HMI tags "BWTS_BTCS"
   "80_From_HMI_RUN_BTCS" : Bool = PLC "80_From_HMI".RUN_BTCS, 1 s
   "80_From_HMI_RUN_BWTS" : Bool = PLC "80_From_HMI".RUN_BWTS, 1 s
   "2110_BTCS_CNTRL_DB_PRE_DWELL_HRS" : Int = PLC "2110_BTCS_CNTRL_DB".PRE_DWELL_HRS, 1 s
   "2110_BTCS_CNTRL_DB_DE_OX_HRS" : Int = PLC "80_From_HMI".MAN_AQ_INC_96, 1 s
   "2110_BTCS_CNTRL_DB_DE_OX_SP_HRS" : Int = PLC "2110_BTCS_CNTRL_DB".DE_OX_SP_HRS, 1 s
   "2110_BTCS_CNTRL_DB_DWELL_HRS" : Int = PLC "2110_BTCS_CNTRL_DB".DWELL_HRS, 1 s
   "2110_BTCS_CNTRL_DB_RE_OX_HRS" : Int = PLC "2110_BTCS_CNTRL_DB".RE_OX_HRS, 1 s
   "2110_BTCS_CNTRL_DB_RE_OX_SP_HRS" : Int = PLC "2110_BTCS_CNTRL_DB".RE_OX_SP_HRS, 1 s
   "2110_BTCS_CNTRL_DB_POST_DWELL_HRS" : Int = PLC "2110_BTCS_CNTRL_DB".POST_DWELL_HRS, 1 s
   "2110_BTCS_CNTRL_DB_PRE_DWELL_MINS" : Int = PLC "2110_BTCS_CNTRL_DB".PRE_DWELL_MINS, 1 s
   "2110_BTCS_CNTRL_DB_DE_OX_MINS" : Int = PLC "2110_BTCS_CNTRL_DB".DE_OX_MINS, 1 s
   "2110_BTCS_CNTRL_DB_DE_OX_SP_MINS" : Int = PLC "2110_BTCS_CNTRL_DB".DE_OX_SP_MINS, 1 s
   "2110_BTCS_CNTRL_DB_DWELL_MINS" : Int = PLC "2110_BTCS_CNTRL_DB".DWELL_MINS, 1 s
   "2110_BTCS_CNTRL_DB_RE_OX_MINS" : Int = PLC "2110_BTCS_CNTRL_DB".RE_OX_MINS, 1 s
   "2110_BTCS_CNTRL_DB_RE_OX_SP_MINS" : Int = PLC "2110_BTCS_CNTRL_DB".RE_OX_SP_MINS, 1 s
   "2110_BTCS_CNTRL_DB_POST_DWELL_MINS" : Int = PLC "2110_BTCS_CNTRL_DB".POST_DWELL_MINS, 1 s
   "2110_BTCS_CNTRL_DB_TOT_SEQ_HRS" : Int = PLC "2110_BTCS_CNTRL_DB".TOT_SEQ_HRS, 1 s
   "2110_BTCS_CNTRL_DB_TOT_SEQ_MINS" : Int = PLC "2110_BTCS_CNTRL_DB".TOT_SEQ_MINS, 1 s
   "2110_BTCS_CNTRL_DB_RMNG_SEQ_HRS" : Int = PLC "84_Setpoints".PIT358_InitialFill_Low, 1 s
   "2110_BTCS_CNTRL_DB_RMNG_SEQ_MINS" : Int = PLC "2110_BTCS_CNTRL_DB".RMNG_SEQ_MINS, 1 s
   "2110_BTCS_CNTRL_DB_BTCS_STATE" : Int = PLC "2110_BTCS_CNTRL_DB".BTCS_STATE, 1 s
   "2110_BTCS_CNTRL_DB_BTCS_STEP" : Int = PLC "2110_BTCS_CNTRL_DB".BTCS_STEP, 1 s
   "2110_BTCS_CNTRL_DB_START_SEQ" : Bool = PLC "2110_BTCS_CNTRL_DB".START_SEQ, 1 s
   "2110_BTCS_CNTRL_DB_STOP_SEQ" : Bool = PLC "2110_BTCS_CNTRL_DB".STOP_SEQ, 1 s
   "2102_TIME_CALCS_DB_TIMES_VALID" : Bool = PLC "2102_TIME_CALCS_DB".TIMES_VALID, 1 s
   "2110_BTCS_CNTRL_DB_PORT_TANK_STS" : Bool = PLC "2110_BTCS_CNTRL_DB".PORT_TANK_STS, 1 s
   "2110_BTCS_CNTRL_DB_RESET_ALL" : Bool = PLC "2110_BTCS_CNTRL_DB".RESET_ALL, 1 s
   "2110_BTCS_CNTRL_DB_STBD_TANK_STS" : Bool = PLC "2110_BTCS_CNTRL_DB".STBD_TANK_STS, 1 s
   "20_TANKS_IP_DATA_RIO_02_FIRST_TANK_BWT_DO" : Real = PLC "20_TANKS_IP_DATA".RIO_02.FIRST_TANK.BWT_DO, 1 s
   "20_TANKS_IP_DATA_RIO_02_FIRST_TANK_BWT_LEVEL" : Real = PLC "20_TANKS_IP_DATA".RIO_02.FIRST_TANK.BWT_LEVEL, 1 s
   "20_TANKS_IP_DATA_RIO_02_FIRST_TANK_BWT_PH" : Real = PLC "20_TANKS_IP_DATA".RIO_02.FIRST_TANK.BWT_PH, 1 s
   "20_TANKS_IP_DATA_RIO_02_FIRST_TANK_BWT_TEMP" : Real = PLC "20_TANKS_IP_DATA".RIO_02.FIRST_TANK.BWT_TEMP, 1 s
   "20_TANKS_IP_DATA_RIO_02_SECOND_TANK_BWT_DO" : Real = PLC "20_TANKS_IP_DATA".RIO_02.SECOND_TANK.BWT_DO, 1 s
   "20_TANKS_IP_DATA_RIO_02_SECOND_TANK_BWT_LEVEL" : Real = PLC "20_TANKS_IP_DATA".RIO_02.SECOND_TANK.BWT_LEVEL, 1 s
   "20_TANKS_IP_DATA_RIO_02_SECOND_TANK_BWT_PH" : Real = PLC "20_TANKS_IP_DATA".RIO_02.SECOND_TANK.BWT_PH, 1 s
   "20_TANKS_IP_DATA_RIO_02_SECOND_TANK_BWT_TEMP" : Real = PLC "20_TANKS_IP_DATA".RIO_02.SECOND_TANK.BWT_TEMP, 1 s
   "2100_AUTO_SEQ_DB_SEQ_RNG" : Bool = PLC "2100_AUTO_SEQ_DB".SEQ_RNG, 1 s
   "2102_TIME_CALCS_DB_POST_DWELL_MINS_RMNG" : Int = PLC "2102_TIME_CALCS_DB".POST_DWELL_MINS_RMNG, 1 s
   "2102_TIME_CALCS_DB_RE_OX_SP_MINS_RMNG" : Int = PLC "2102_TIME_CALCS_DB".RE_OX_SP_MINS_RMNG, 1 s
   "2102_TIME_CALCS_DB_RE_OX_MINS_RMNG" : Int = PLC "2102_TIME_CALCS_DB".RE_OX_MINS_RMNG, 1 s
   "2102_TIME_CALCS_DB_DE_OX_SP_MINS_RMNG" : Int = PLC "2102_TIME_CALCS_DB".DE_OX_SP_MINS_RMNG, 1 s
   "2102_TIME_CALCS_DB_DWELL_MINS_RMNG" : Int = PLC "2102_TIME_CALCS_DB".DWELL_MINS_RMNG, 1 s
   "2102_TIME_CALCS_DB_DE_OX_MINS_RMNG" : Int = PLC "2102_TIME_CALCS_DB".DE_OX_MINS_RMNG, 1 s
   "2102_TIME_CALCS_DB_PRE_DWELL_MINS_RMNG" : Int = PLC "2102_TIME_CALCS_DB".PRE_DWELL_MINS_RMNG, 1 s
   "2102_TIME_CALCS_DB_RE_OX_SP_TMR_DN" : Bool = PLC "2102_TIME_CALCS_DB".RE_OX_SP_TMR_DN, 1 s
   "2102_TIME_CALCS_DB_DE_OX_SP_TMR_DN" : Bool = PLC "2102_TIME_CALCS_DB".DE_OX_SP_TMR_DN, 1 s
   "2102_TIME_CALCS_DB_DWELL_TMR_DN" : Bool = PLC "2102_TIME_CALCS_DB".DWELL_TMR_DN, 1 s
   "2102_TIME_CALCS_DB_POST_DWELL_TMR_DN" : Bool = PLC "2102_TIME_CALCS_DB".POST_DWELL_TMR_DN, 1 s
   "2102_TIME_CALCS_DB_DE_OX_TMR_DN" : Bool = PLC "2102_TIME_CALCS_DB".DE_OX_TMR_DN, 1 s
   "2102_TIME_CALCS_DB_PRE_DWELL_TMR_DN" : Bool = PLC "2102_TIME_CALCS_DB".PRE_DWELL_TMR_DN, 1 s
   "2102_TIME_CALCS_DB_TOT_SEQ_MINS_RMNG" : Int = PLC "2102_TIME_CALCS_DB".TOT_SEQ_MINS_RMNG, 1 s
   "2102_TIME_CALCS_DB_TOT_SEQ_HRS_RMNG" : Int = PLC "2102_TIME_CALCS_DB".TOT_SEQ_HRS_RMNG, 1 s
   "2102_TIME_CALCS_DB_RE_OX_TMR_DN" : Bool = PLC "2102_TIME_CALCS_DB".RE_OX_TMR_DN, 1 s
   "1405_PID_CV405_CtrlParamsBackUp_Gain" : Real = PLC "1405_PID_CV405".CtrlParamsBackUp.Gain, 1 s
   "1405_PID_CV405_CtrlParamsBackUp_Ti" : Real = PLC "1405_PID_CV405".CtrlParamsBackUp.Ti, 1 s
   "20_TANKS_IP_DATA_RIO_02_FIRST_TANK_TANK_VENT_A_OPEN" : Bool = PLC "20_TANKS_IP_DATA".RIO_02.FIRST_TANK.TANK_VENT_A_OPEN AT %DB1.DBW0, 1 s
   "40_TANKS_OP_DATA_RIO_02_VENT_A_2P" : Bool = PLC "40_TANKS_OP_DATA".RIO_02_VENT_A_2P AT %DB1.DBW0, 1 s
   "20_TANKS_IP_DATA_RIO_02_FIRST_TANK_GTT_ISOL_VALVE_OPEN" : Bool = PLC "20_TANKS_IP_DATA".RIO_02.FIRST_TANK.GTT_ISOL_VALVE_OPEN AT %DB1.DBW0, 1 s
   "20_TANKS_IP_DATA_RIO_02_FIRST_TANK_GTT_ISOL_VALVE_CLSD" : Bool = PLC "20_TANKS_IP_DATA".RIO_02.FIRST_TANK.GTT_ISOL_VALVE_CLSD AT %DB1.DBW0, 1 s
   "20_TANKS_IP_DATA_RIO_02_FIRST_TANK_TANK_VENT_A_CLSD" : Bool = PLC "20_TANKS_IP_DATA".RIO_02.FIRST_TANK.TANK_VENT_A_CLSD AT %DB1.DBW0, 1 s
   "40_TANKS_OP_DATA_RIO_02_VENT_B_2P" : Bool = PLC "40_TANKS_OP_DATA".RIO_02_VENT_B_2P AT %DB1.DBW0, 1 s
   "20_TANKS_IP_DATA_RIO_02_FIRST_TANK_TANK_VENT_B_OPEN" : Bool = PLC "20_TANKS_IP_DATA".RIO_02.FIRST_TANK.TANK_VENT_B_OPEN AT %DB1.DBW0, 1 s
   "20_TANKS_IP_DATA_RIO_02_FIRST_TANK_TANK_VENT_B_CLSD" : Bool = PLC "20_TANKS_IP_DATA".RIO_02.FIRST_TANK.TANK_VENT_B_CLSD AT %DB1.DBW0, 1 s
   "40_TANKS_OP_DATA_RIO_02_VENT_B_2P(1)" : Bool = PLC "40_TANKS_OP_DATA".RIO_02_VENT_B_2P AT %DB1.DBW0, 1 s
   "20_TANKS_IP_DATA_RIO_02_SECOND_TANK_TANK_VENT_B_OPEN" : Bool = PLC "20_TANKS_IP_DATA".RIO_02.SECOND_TANK.TANK_VENT_B_OPEN AT %DB1.DBW0, 1 s
   "20_TANKS_IP_DATA_RIO_02_SECOND_TANK_TANK_VENT_B_CLSD" : Bool = PLC "20_TANKS_IP_DATA".RIO_02.SECOND_TANK.TANK_VENT_B_CLSD AT %DB1.DBW0, 1 s
   "40_TANKS_OP_DATA_RIO_02_VENT_B_2S(1)" : Bool = PLC "40_TANKS_OP_DATA".RIO_02_VENT_B_2S AT %DB1.DBW0, 1 s
   "20_TANKS_IP_DATA_RIO_02_SECOND_TANK_TANK_VENT_A_OPEN" : Bool = PLC "20_TANKS_IP_DATA".RIO_02.SECOND_TANK.TANK_VENT_A_OPEN AT %DB1.DBW0, 1 s
   "20_TANKS_IP_DATA_RIO_02_SECOND_TANK_TANK_VENT_A_CLSD" : Bool = PLC "20_TANKS_IP_DATA".RIO_02.SECOND_TANK.TANK_VENT_A_CLSD AT %DB1.DBW0, 1 s
   "20_TANKS_IP_DATA_RIO_02_FIRST_TANK_BWT_LEVEL_HIHI" : Bool = PLC "20_TANKS_IP_DATA".RIO_02.FIRST_TANK.BWT_LEVEL_HIHI AT %DB1.DBW0, 1 s
   "20_TANKS_IP_DATA_RIO_02_SECOND_TANK_BWT_LEVEL_HIHI" : Bool = PLC "20_TANKS_IP_DATA".RIO_02.SECOND_TANK.BWT_LEVEL_HIHI AT %DB1.DBW0, 1 s
   "20_TANKS_IP_DATA_RIO_02_FIRST_TANK_TANKS_PRESS_HIHI" : Bool = PLC "20_TANKS_IP_DATA".RIO_02.FIRST_TANK.TANKS_PRESS_HIHI AT %DB1.DBW0, 1 s
   "20_TANKS_IP_DATA_RIO_02_SECOND_TANK_TANKS_PRESS_HIHI" : Bool = PLC "20_TANKS_IP_DATA".RIO_02.SECOND_TANK.TANKS_PRESS_HIHI AT %DB1.DBW0, 1 s
   "20_TANKS_IP_DATA_RIO_02_FIRST_TANK_TANKS_PRESS" : Real = PLC "20_TANKS_IP_DATA".RIO_02.FIRST_TANK.TANKS_PRESS AT %DB1.DBW0, 1 s
   "20_TANKS_IP_DATA_RIO_02_FIRST_TANK_USD_FLOW" : Real = PLC "20_TANKS_IP_DATA".RIO_02.FIRST_TANK.USD_FLOW AT %DB1.DBW0, 1 s
   "20_TANKS_IP_DATA_RIO_02_FIRST_TANK_MBG_FLOW" : Real = PLC "20_TANKS_IP_DATA".RIO_02.FIRST_TANK.MBG_FLOW AT %DB1.DBW0, 1 s
   "20_TANKS_IP_DATA_RIO_02_FIRST_TANK_O2_MONITOR" : Real = PLC "20_TANKS_IP_DATA".RIO_02.FIRST_TANK.O2_MONITOR AT %DB1.DBW0, 1 s
   "20_TANKS_IP_DATA_RIO_02_SECOND_TANK_TANKS_PRESS" : Real = PLC "20_TANKS_IP_DATA".RIO_02.SECOND_TANK.TANKS_PRESS AT %DB1.DBW0, 1 s
   "20_TANKS_IP_DATA_RIO_02_SECOND_TANK_USD_FLOW" : Real = PLC "20_TANKS_IP_DATA".RIO_02.SECOND_TANK.USD_FLOW AT %DB1.DBW0, 1 s
   "20_TANKS_IP_DATA_RIO_02_SECOND_TANK_MBG_FLOW" : Real = PLC "20_TANKS_IP_DATA".RIO_02.SECOND_TANK.MBG_FLOW AT %DB1.DBW0, 1 s
   "20_TANKS_IP_DATA_RIO_02_SECOND_TANK_O2_MONITOR" : Real = PLC "20_TANKS_IP_DATA".RIO_02.SECOND_TANK.O2_MONITOR AT %DB1.DBW0, 1 s
   "20_TANKS_IP_DATA_RIO_02_SECOND_TANK_DECK_IG_PRESS" : Real = PLC "20_TANKS_IP_DATA".RIO_02.SECOND_TANK.DECK_IG_PRESS AT %DB1.DBW0, 1 s
   "20_TANKS_IP_DATA_RIO_02_SECOND_TANK_GTT_ISOL_VALVE_OPEN" : Bool = PLC "20_TANKS_IP_DATA".RIO_02.SECOND_TANK.GTT_ISOL_VALVE_OPEN AT %DB1.DBW0, 1 s
   "20_TANKS_IP_DATA_RIO_02_SECOND_TANK_GTT_ISOL_VALVE_CLSD" : Bool = PLC "20_TANKS_IP_DATA".RIO_02.SECOND_TANK.GTT_ISOL_VALVE_CLSD AT %DB1.DBW0, 1 s
   "2019_AUT_MAN_CNTRL_PORT_GTT_VLV_MAN" : Bool = PLC "2019_AUT_MAN_CNTRL".PORT_GTT_VLV_MAN AT %DB1.DBW0, 1 s
   "2019_AUT_MAN_CNTRL_STBD_GTT_VLV_MAN" : Bool = PLC "2019_AUT_MAN_CNTRL".STBD_GTT_VLV_MAN AT %DB1.DBW0, 1 s
   "14_DQ_DATA_CV_422_2P" : Bool = PLC "14_DQ_DATA".CV_422_2P AT %DB1.DBW0, 1 s
   "14_DQ_DATA_CV_421_2S" : Bool = PLC "14_DQ_DATA".CV_421_2S AT %DB1.DBW0, 1 s
   "2086_Times_DEOX_PRE_GTT_OPN_DLY" : Time = PLC "2086_Times".DEOX_PRE_GTT_OPN_DLY AT %DB1.DBW0, 1 s
   "2086_Times_DEOX_PRE_GTT_CLS_DLY" : Time = PLC "2086_Times".DEOX_PRE_GTT_CLS_DLY AT %DB1.DBW0, 1 s
   "2086_Times_REOX_PRE_GTT_OPN_DLY" : Time = PLC "2086_Times".REOX_PRE_GTT_OPN_DLY AT %DB1.DBW0, 1 s
   "2086_Times_REOX_PRE_GTT_CLS_DLY" : Time = PLC "2086_Times".REOX_PRE_GTT_CLS_DLY AT %DB1.DBW0, 1 s
   "2086_Times_AT_DEOX_CNF_TIME" : Time = PLC "2086_Times".AT_DEOX_CNF_TIME AT %DB1.DBW0, 1 s
   "2086_Times_AT_REOX_CNF_TIME" : Time = PLC "2086_Times".AT_REOX_CNF_TIME AT %DB1.DBW0, 1 s
   "2084_Setpoints_FIT418_LoLo" : Real = PLC "2084_Setpoints".FIT418_LoLo AT %DB1.DBW0, 1 s
   "2084_Setpoints_PIT424_HiHi" : Real = PLC "2084_Setpoints".PIT424_HiHi AT %DB1.DBW0, 1 s
   "2084_Setpoints_PIT424_Hi" : Real = PLC "2084_Setpoints".PIT424_Hi AT %DB1.DBW0, 1 s
   "2084_Setpoints_PIT424_Lo" : Real = PLC "2084_Setpoints".PIT424_Lo AT %DB1.DBW0, 1 s
   "2084_Setpoints_PIT424_LoLo" : Real = PLC "2084_Setpoints".PIT424_LoLo AT %DB1.DBW0, 1 s
   "2084_Setpoints_PIT415_HiHi" : Real = PLC "2084_Setpoints".PIT415_HiHi AT %DB1.DBW0, 1 s
   "2084_Setpoints_PIT415_Hi" : Real = PLC "2084_Setpoints".PIT415_Hi AT %DB1.DBW0, 1 s
   "2084_Setpoints_PIT415_Lo" : Real = PLC "2084_Setpoints".PIT415_Lo AT %DB1.DBW0, 1 s
   "2084_Setpoints_PIT415_LoLo" : Real = PLC "2084_Setpoints".PIT415_LoLo AT %DB1.DBW0, 1 s
   "2084_Setpoints_DO_SP" : Real = PLC "2084_Setpoints".DO_SP AT %DB1.DBW0, 1 s
   "2084_Setpoints_TT436_Hi" : Real = PLC "2084_Setpoints".TT436_Hi AT %DB1.DBW0, 1 s
   "2084_Setpoints_LT422_Hi" : Real = PLC "2084_Setpoints".LT422_Hi AT %DB1.DBW0, 1 s
   "2084_Setpoints_LT422_Lo" : Real = PLC "2084_Setpoints".LT422_Lo AT %DB1.DBW0, 1 s
   "2084_Setpoints_FIT420_HiHi" : Real = PLC "2084_Setpoints".FIT420_HiHi AT %DB1.DBW0, 1 s
   "2084_Setpoints_FIT420_Hi" : Real = PLC "2084_Setpoints".FIT420_Hi AT %DB1.DBW0, 1 s
   "2084_Setpoints_FIT420_Lo" : Real = PLC "86_Times".PIT402_Ramp_Seconds AT %DB1.DBW0, 1 s
   "2084_Setpoints_FIT420_LoLo" : Real = PLC "2084_Setpoints".FIT420_LoLo AT %DB1.DBW0, 1 s
   "2084_Setpoints_FIT418_HiHi" : Real = PLC "2084_Setpoints".FIT418_HiHi AT %DB1.DBW0, 1 s
   "2084_Setpoints_PH_SP" : Real = PLC "2084_Setpoints".PH_SP AT %DB1.DBW0, 1 s
   "2084_Setpoints_TT436_HiHi" : Real = PLC "2084_Setpoints".TT436_HiHi AT %DB1.DBW0, 1 s
   "2084_Setpoints_FIT418_Lo" : Real = PLC "2084_Setpoints".FIT418_Lo AT %DB1.DBW0, 1 s
   "2084_Setpoints_FIT418_Hi" : Real = PLC "2084_Setpoints".FIT418_Hi AT %DB1.DBW0, 1 s
   "80_From_HMI_SAL_VALUE" : Real = PLC "80_From_HMI".SAL_VALUE, 1 s
   "80_From_HMI_SAL_CNFRM" : Bool = PLC "80_From_HMI".SAL_CNFRM, 1 s
   "2068_Sys_Status_Data_SAL_VALID" : Bool = PLC "2068_Sys_Status_Data".SAL_VALID, 1 s
   "150_GCU_LCL_CNTRL_DB_OPN_ACTV_GTT_VLVS" : Bool = PLC "150_GCU_LCL_CNTRL_DB".OPN_ACTV_GTT_VLVS, 1 s
   "80_From_HMI_LOW_SAL_ACPT" : Bool = PLC "80_From_HMI".LOW_SAL_ACPT, 1 s
   "80_From_HMI_LOW_SAL_RJCT" : Bool = PLC "80_From_HMI".LOW_SAL_RJCT, 1 s
   "2068_Sys_Status_Data_SAL_CNF_CHK" : Bool = PLC "2068_Sys_Status_Data".SAL_CNF_CHK, 100 ms
      on ChangeValue: "Salinity_FreshWaterAlert"()
   "20_TANKS_IP_DATA_RIO_02_FIRST_TANK_USD FLOW  N" : Real = PLC "20_TANKS_IP_DATA".RIO_02.FIRST_TANK."USD FLOW  N" AT %DB1.DBD0, 1 s
   "20_TANKS_IP_DATA_RIO_02_FIRST_TANK_MBG_FLOW N" : Real = PLC "20_TANKS_IP_DATA".RIO_02.FIRST_TANK."MBG_FLOW N" AT %DB1.DBD0, 1 s
   "20_TANKS_IP_DATA_RIO_02_SECOND_TANK_MBG_FLOW N" : Real = PLC "20_TANKS_IP_DATA".RIO_02.SECOND_TANK."MBG_FLOW N" AT %DB1.DBD0, 1 s
   "20_TANKS_IP_DATA_RIO_02_SECOND_TANK_USD FLOW  N" : Real = PLC "20_TANKS_IP_DATA".RIO_02.SECOND_TANK."USD FLOW  N" AT %DB1.DBD0, 1 s

HMI tags "GCU"
   "10_DI_DATA_P_303_ENBLD" : Bool = PLC "10_DI_DATA".P_303_ENBLD, 1 s
   "10_DI_DATA_P_304_ENBLD" : Bool = PLC "10_DI_DATA".P_304_ENBLD, 1 s
   "12_AI_Data_CV_405_SCALED" : Real = PLC "12_AI_Data".CV_405_SCALED, 1 s
   "10_DI_DATA_P_303_OK" : Bool = PLC "10_DI_DATA".P_303_OK, 1 s
   "10_DI_DATA_P_304_OK" : Bool = PLC "10_DI_DATA".P_304_OK, 1 s
   "16_AQ_Data_CV405_CNTRL" : Real = PLC "16_AQ_Data".CV405_CNTRL, 1 s
   "10_DI_DATA_CV358_CLSD" : Bool = PLC "10_DI_DATA".CV358_CLSD, 1 s
   "10_DI_DATA_E_400_RUN" : Bool = PLC "10_DI_DATA".E_400_RUN, 1 s
   "10_DI_DATA_CV341_CLSD" : Bool = PLC "10_DI_DATA".CV341_CLSD, 1 s
   "10_DI_DATA_CV341_OPN" : Bool = PLC "10_DI_DATA".CV341_OPN, 1 s
   "10_DI_DATA_CV411_CLSD" : Bool = PLC "10_DI_DATA".CV411_CLSD, 1 s
   "10_DI_DATA_CV411_OPN" : Bool = PLC "10_DI_DATA".CV411_OPN, 1 s
   "10_DI_DATA_CV407_OPN" : Bool = PLC "10_DI_DATA".CV407_OPN, 1 s
   "10_DI_DATA_CV409_CLSD" : Bool = PLC "10_DI_DATA".CV409_CLSD, 1 s
   "10_DI_DATA_CV409_OPN" : Bool = PLC "10_DI_DATA".CV409_OPN, 1 s
   "10_DI_DATA_CV406_OPN" : Bool = PLC "10_DI_DATA".CV406_OPN, 1 s
   "10_DI_DATA_FS_350_FLW_OK" : Bool = PLC "10_DI_DATA".FS_350_FLW_OK, 1 s
   "12_AI_Data_LIT_304_SCALED" : Real = PLC "12_AI_Data".LIT_304_SCALED, 1 s
   "10_DI_DATA_FS_332 FLW_OK" : Bool = PLC "10_DI_DATA"."FS_332 FLW_OK", 1 s
   "10_DI_DATA_CV406_CLSD" : Bool = PLC "10_DI_DATA".CV406_CLSD, 1 s
   "10_DI_DATA_CV407_CLSD" : Bool = PLC "10_DI_DATA".CV407_CLSD, 1 s
   "12_AI_Data_E_400_PT002_SCALED" : Real = PLC "12_AI_Data".E_400_PT002_SCALED, 1 s
   "12_AI_Data_TIT_406_SCALED" : Real = PLC "12_AI_Data".TIT_406_SCALED, 1 s
   "12_AI_Data_PIT_416_SCALED" : Real = PLC "12_AI_Data".PIT_416_SCALED, 1 s
   "12_AI_Data_PIT_353_SCALED" : Real = PLC "12_AI_Data".PIT_353_SCALED, 1 s
   "12_AI_Data_TIT_408_SCALED" : Real = PLC "12_AI_Data".TIT_408_SCALED, 1 s
   "12_AI_Data_PIT_348_SCALED" : Real = PLC "12_AI_Data".PIT_348_SCALED, 1 s
   "12_AI_Data_PIT_358_SCALED" : Real = PLC "12_AI_Data".PIT_358_SCALED, 1 s
   "12_AI_Data_E_400_TE002_SCALED" : Real = PLC "12_AI_Data".E_400_TE002_SCALED, 1 s
   "10_DI_DATA_LS_303_LO" : Bool = PLC "10_DI_DATA".LS_303_LO, 1 s
   "10_DI_DATA_CV441_CLSD" : Bool = PLC "10_DI_DATA".CV441_CLSD, 1 s
   "10_DI_DATA_CV441_OPN" : Bool = PLC "10_DI_DATA".CV441_OPN, 1 s
   "20_TANKS_IP_DATA_RIO_02_FIRST_TANK_DECK_IG_PRESS" : Real = PLC "20_TANKS_IP_DATA".RIO_02.FIRST_TANK.DECK_IG_PRESS, 1 s
   "10_DI_DATA_CV358_OPN" : Bool = PLC "10_DI_DATA".CV358_OPN, 1 s
   "84_Setpoints_LIT304_InitialFill_High" : Real = PLC "84_Setpoints".LIT304_InitialFill_High, 1 s
   "84_Setpoints_LIT304_InitialFill_Low" : Real = PLC "84_Setpoints".LIT304_InitialFill_Low, 1 s
   "10_DI_DATA_E_400_NOK" : Bool = PLC "10_DI_DATA".E_400_NOK, 1 s
   "10_DI_DATA_E_400_SHTDN" : Bool = PLC "10_DI_DATA".E_400_SHTDN, 1 s
   "140_PGC_HRS_RUN_DB_RST" : Bool = PLC "140_PGC_HRS_RUN_DB".RST, 1 s
   "140_PGC_HRS_RUN_DB_SRVC" : Bool = PLC "140_PGC_HRS_RUN_DB".SRVC, 1 s
   "140_PGC_HRS_RUN_DB_SECS" : Int = PLC "140_PGC_HRS_RUN_DB".SECS, 1 s
   "140_PGC_HRS_RUN_DB_MINS" : Int = PLC "140_PGC_HRS_RUN_DB".MINS, 1 s
   "140_PGC_HRS_RUN_DB_HRS" : Int = PLC "140_PGC_HRS_RUN_DB".HRS, 1 s
   "140_PGC_HRS_RUN_DB_SRV_HRS" : Int = PLC "140_PGC_HRS_RUN_DB".SRV_HRS, 1 s
   "140_PGC_HRS_RUN_DB_SHRS_IP" : Int = PLC "140_PGC_HRS_RUN_DB".SHRS_IP, 1 s
   "84_Setpoints_E400_TT002_HighHigh" : Real = PLC "84_Setpoints".E400_TT002_HighHigh, 1 s
   "84_Setpoints_E400_PT002_HighHigh" : Real = PLC "84_Setpoints".E400_PT002_HighHigh, 1 s
   "19_AUTO_CMNDS_Data_CV405_PID_MDLTG" : Bool = PLC "19_AUTO_CMNDS_Data".CV405_PID_MDLTG, 1 s
   "84_Setpoints_PIT416_HighHigh" : Real = PLC "84_Setpoints".PIT416_HighHigh, 1 s
   "12_AI_Data_R3_SPR_AI_802_SCALED" : Real = PLC "12_AI_Data".R3_SPR_AI_802_SCALED, 1 s
   "12_AI_Data_R3_SPR_AI_824_SCALED" : Real = PLC "12_AI_Data".R3_SPR_AI_824_SCALED, 1 s
   "12_AI_Data_R3_SPR_AI_826_SCALED" : Real = PLC "12_AI_Data".R3_SPR_AI_826_SCALED, 1 s
   "12_AI_Data_R3_SPR_AI_828_SCALED" : Real = PLC "12_AI_Data".R3_SPR_AI_828_SCALED, 1 s
   "12_AI_Data_R3_SPR_AI_830_SCALED" : Real = PLC "12_AI_Data".R3_SPR_AI_830_SCALED, 1 s
   "12_AI_Data_SL_400_SCALED" : Real = PLC "12_AI_Data".SL_400_SCALED, 1 s
   "10_DI_DATA_5T1_PWR_OK" : Bool = PLC "10_DI_DATA".5T1_PWR_OK, 1 s
   "10_DI_DATA_6Q6_PWR_OK" : Bool = PLC "10_DI_DATA".6Q6_PWR_OK, 1 s
   "19_AUTO_CMNDS_Data_PIT353_CMND_LowLow" : Real = PLC "19_AUTO_CMNDS_Data".PIT353_CMND_LowLow, 1 s
   "19_AUTO_CMNDS_Data_PIT353_CMND_Low" : Real = PLC "19_AUTO_CMNDS_Data".PIT353_CMND_Low, 1 s
   "84_Setpoints_TIT408_High" : Real = PLC "84_Setpoints".TIT408_High, 1 s
   "10_DI_DATA_PB_10S1" : Bool = PLC "10_DI_DATA".PB_10S1, 1 s
   "10_DI_DATA_PB_10S2" : Bool = PLC "10_DI_DATA".PB_10S2, 1 s
   "10_DI_DATA_EPB_8S1" : Bool = PLC "10_DI_DATA".EPB_8S1, 1 s
   "10_DI_DATA_E_400_STPD" : Bool = PLC "10_DI_DATA".E_400_STPD, 1 s
   "10_DI_DATA_R3_SPR_DI_136_1" : Bool = PLC "10_DI_DATA".R3_SPR_DI_136_1, 1 s
   "10_DI_DATA_R3_SPR_DI_136_0" : Bool = PLC "10_DI_DATA".R3_SPR_DI_136_0, 1 s
   "19_AUTO_CMNDS_Data_LIT304_CMND_HighHigh" : Real = PLC "19_AUTO_CMNDS_Data".LIT304_CMND_HighHigh, 1 s
   "19_AUTO_CMNDS_Data_LIT304_CMND_Target" : Real = PLC "19_AUTO_CMNDS_Data".LIT304_CMND_Target, 1 s
   "19_AUTO_CMNDS_Data_PIT353_CMND_High" : Real = PLC "19_AUTO_CMNDS_Data".PIT353_CMND_High, 1 s
   "19_AUTO_CMNDS_Data_PIT353_CMND_HighHigh" : Real = PLC "19_AUTO_CMNDS_Data".PIT353_CMND_HighHigh, 1 s
   "84_Setpoints_E400_PT002_High" : Real = PLC "84_Setpoints".E400_PT002_High, 1 s
   "84_Setpoints_E400_TT002_High" : Real = PLC "84_Setpoints".E400_TT002_High, 1 s
   "84_Setpoints_PIT348_LowLow" : Real = PLC "84_Setpoints".PIT348_LowLow, 1 s
   "84_Setpoints_PIT348_Low" : Real = PLC "84_Setpoints".PIT348_Low, 1 s
   "84_Setpoints_PIT348_High" : Real = PLC "84_Setpoints".PIT348_High, 1 s
   "84_Setpoints_PIT348_HighHigh" : Real = PLC "84_Setpoints".PIT348_HighHigh, 1 s
   "19_AUTO_CMNDS_Data_PIT358_CMND_Low" : Real = PLC "19_AUTO_CMNDS_Data".PIT358_CMND_Low, 1 s
   "19_AUTO_CMNDS_Data_PIT358_CMND_LowLow" : Real = PLC "19_AUTO_CMNDS_Data".PIT358_CMND_LowLow, 1 s
   "19_AUTO_CMNDS_Data_PIT358_CMND_High" : Real = PLC "19_AUTO_CMNDS_Data".PIT358_CMND_High, 1 s
   "84_Setpoints_PIT416_LowLow" : Real = PLC "84_Setpoints".PIT416_LowLow, 1 s
   "84_Setpoints_PIT416_Low" : Real = PLC "84_Setpoints".PIT416_Low, 1 s
   "84_Setpoints_PIT416_Target" : Real = PLC "84_Setpoints".PIT416_Target, 1 s
   "84_Setpoints_PIT416_High" : Real = PLC "84_Setpoints".PIT416_High, 1 s
   "84_Setpoints_TIT408_HighHigh" : Real = PLC "84_Setpoints".TIT408_HighHigh, 1 s
   "84_Setpoints_TIT406_High" : Real = PLC "84_Setpoints".TIT406_High, 1 s
   "84_Setpoints_TIT406_HighHigh" : Real = PLC "84_Setpoints".TIT406_HighHigh, 1 s
   "19_AUTO_CMNDS_Data_LIT304_CMND_LowLow" : Real = PLC "19_AUTO_CMNDS_Data".LIT304_CMND_LowLow, 1 s
   "19_AUTO_CMNDS_Data_LIT304_CMND_High" : Real = PLC "19_AUTO_CMNDS_Data".LIT304_CMND_High, 1 s
   "19_AUTO_CMNDS_Data_LIT304_CMND_Low" : Real = PLC "19_AUTO_CMNDS_Data".LIT304_CMND_Low, 1 s
   "19_AUTO_CMNDS_Data_PIT358_CMND_HighHigh" : Real = PLC "19_AUTO_CMNDS_Data".PIT358_CMND_HighHigh, 1 s
   "84_Setpoints_LIT304_InitialFill_Target" : Real = PLC "84_Setpoints".LIT304_InitialFill_Target, 1 s
   "84_Setpoints_LIT304_InitialFill_HighHigh" : Real = PLC "84_Setpoints".LIT304_InitialFill_HighHigh, 1 s
   "84_Setpoints_LIT304_InitialFill_LowLow" : Real = PLC "84_Setpoints".LIT304_InitialFill_LowLow, 1 s
   "84_Setpoints_LIT304_Refill_HighHigh" : Real = PLC "84_Setpoints".LIT304_Refill_HighHigh, 1 s
   "84_Setpoints_LIT304_Refill_Target" : Real = PLC "84_Setpoints".LIT304_Refill_Target, 1 s
   "84_Setpoints_LIT304_Refill_Low" : Real = PLC "84_Setpoints".LIT304_Refill_Low, 1 s
   "84_Setpoints_LIT304_Refill_LowLow" : Real = PLC "84_Setpoints".LIT304_Refill_LowLow, 1 s
   "84_Setpoints_LIT304_Refill_High" : Real = PLC "84_Setpoints".LIT304_Refill_High, 1 s
   "84_Setpoints_PIT358_InitialFill_LowLow" : Real = PLC "84_Setpoints".PIT358_InitialFill_LowLow, 1 s
   "84_Setpoints_PIT358_InitialFill_Low" : Real = PLC "84_Setpoints".PIT358_InitialFill_Low, 1 s
   "84_Setpoints_PIT358_InitialFill_High" : Real = PLC "84_Setpoints".PIT358_InitialFill_High, 1 s
   "84_Setpoints_PIT358_InitialFill_HighHigh" : Real = PLC "84_Setpoints".PIT358_InitialFill_HighHigh, 1 s
   "84_Setpoints_PIT358_Refill_LowLow" : Real = PLC "84_Setpoints".PIT358_Refill_LowLow, 1 s
   "84_Setpoints_PIT358_Refill_Low" : Real = PLC "84_Setpoints".PIT358_Refill_Low, 1 s
   "84_Setpoints_PIT358_Refill_High" : Real = PLC "84_Setpoints".PIT358_Refill_High, 1 s
   "84_Setpoints_PIT358_Refill_HighHigh" : Real = PLC "84_Setpoints".PIT358_Refill_HighHigh, 1 s
   "84_Setpoints_PIT353_InitialFill_LowLow" : Real = PLC "84_Setpoints".PIT353_InitialFill_LowLow, 1 s
   "84_Setpoints_PIT353_InitialFill_Low" : Real = PLC "84_Setpoints".PIT353_InitialFill_Low, 1 s
   "84_Setpoints_PIT353_InitialFill_High" : Real = PLC "84_Setpoints".PIT353_InitialFill_High, 1 s
   "84_Setpoints_PIT353_InitialFill_HighHigh" : Real = PLC "84_Setpoints".PIT353_InitialFill_HighHigh, 1 s
   "84_Setpoints_PIT353_Refill_LowLow" : Real = PLC "84_Setpoints".PIT353_Refill_LowLow, 1 s
   "84_Setpoints_PIT353_Refill_Low" : Real = PLC "84_Setpoints".PIT353_Refill_Low, 1 s
   "84_Setpoints_PIT353_Refill_High" : Real = PLC "84_Setpoints".PIT353_Refill_High, 1 s
   "84_Setpoints_PIT353_Refill_HighHigh" : Real = PLC "84_Setpoints".PIT353_Refill_HighHigh, 1 s
   "82_To_HMI_CRNT_MODE_GCU" : Int = PLC "82_To_HMI".CRNT_MODE_GCU, 1 s
   "80_From_HMI_MAN_DQ_136_0" : Bool = PLC "80_From_HMI".MAN_DQ_136_0, 1 s
   "80_From_HMI_MAN_DQ_136_1" : Bool = PLC "80_From_HMI".MAN_DQ_136_1, 1 s
   "80_From_HMI_MAN_DQ_136_2" : Bool = PLC "80_From_HMI".MAN_DQ_136_2, 1 s
   "80_From_HMI_MAN_DQ_136_3" : Bool = PLC "80_From_HMI".MAN_DQ_136_3, 1 s
   "80_From_HMI_MAN_DQ_136_4" : Bool = PLC "80_From_HMI".MAN_DQ_136_4, 1 s
   "80_From_HMI_MAN_DQ_136_5" : Bool = PLC "80_From_HMI".MAN_DQ_136_5, 1 s
   "80_From_HMI_MAN_DQ_136_6" : Bool = PLC "80_From_HMI".MAN_DQ_136_6, 1 s
   "80_From_HMI_MAN_DQ_136_7" : Bool = PLC "80_From_HMI".MAN_DQ_136_7, 1 s
   "80_From_HMI_MAN_DQ_137_0" : Bool = PLC "80_From_HMI".MAN_DQ_137_0, 1 s
   "80_From_HMI_MAN_DQ_137_1" : Bool = PLC "80_From_HMI".MAN_DQ_137_1, 1 s
   "80_From_HMI_MAN_DQ_137_2" : Bool = PLC "80_From_HMI".MAN_DQ_137_2, 1 s
   "80_From_HMI_MAN_DQ_137_3" : Bool = PLC "80_From_HMI".MAN_DQ_137_3, 1 s
   "80_From_HMI_MAN_DQ_137_4" : Bool = PLC "80_From_HMI".MAN_DQ_137_4, 1 s
   "80_From_HMI_MAN_DQ_137_5" : Bool = PLC "80_From_HMI".MAN_DQ_137_5, 1 s
   "80_From_HMI_MAN_DQ_137_6" : Bool = PLC "80_From_HMI".MAN_DQ_137_6, 1 s
   "80_From_HMI_MAN_DQ_137_7" : Bool = PLC "80_From_HMI".MAN_DQ_137_7, 1 s
   "80_From_HMI_MAN_DQ_138_0" : Bool = PLC "80_From_HMI".MAN_DQ_138_0, 1 s
   "80_From_HMI_MAN_DQ_138_1" : Bool = PLC "80_From_HMI".MAN_DQ_138_1, 1 s
   "80_From_HMI_MAN_DQ_138_2" : Bool = PLC "80_From_HMI".MAN_DQ_138_2, 1 s
   "80_From_HMI_MAN_DQ_138_3" : Bool = PLC "80_From_HMI".MAN_DQ_138_3, 1 s
   "80_From_HMI_MAN_DQ_138_4" : Bool = PLC "80_From_HMI".MAN_DQ_138_4, 1 s
   "80_From_HMI_MAN_DQ_138_5" : Bool = PLC "80_From_HMI".MAN_DQ_138_5, 1 s
   "80_From_HMI_MAN_DQ_138_6" : Bool = PLC "80_From_HMI".MAN_DQ_138_6, 1 s
   "80_From_HMI_MAN_DQ_138_7" : Bool = PLC "80_From_HMI".MAN_DQ_138_7, 1 s
   "80_From_HMI_MAN_DQ_139_0" : Bool = PLC "80_From_HMI".MAN_DQ_139_0, 1 s
   "80_From_HMI_MAN_DQ_139_1" : Bool = PLC "80_From_HMI".MAN_DQ_139_1, 1 s
   "80_From_HMI_MAN_DQ_139_2" : Bool = PLC "80_From_HMI".MAN_DQ_139_2, 1 s
   "80_From_HMI_MAN_DQ_139_3" : Bool = PLC "80_From_HMI".MAN_DQ_139_3, 1 s
   "80_From_HMI_MAN_DQ_139_4" : Bool = PLC "80_From_HMI".MAN_DQ_139_4, 1 s
   "80_From_HMI_MAN_DQ_139_5" : Bool = PLC "80_From_HMI".MAN_DQ_139_5, 1 s
   "80_From_HMI_MAN_DQ_139_6" : Bool = PLC "80_From_HMI".MAN_DQ_139_6, 1 s
   "80_From_HMI_MAN_DQ_139_7" : Bool = PLC "80_From_HMI".MAN_DQ_139_7, 1 s
   "16_AQ_Data_R3_SPR_AQ_806" : Real = PLC "16_AQ_Data".R3_SPR_AQ_806, 1 s
   "16_AQ_Data_R3_SPR_AQ_804" : Real = PLC "16_AQ_Data".R3_SPR_AQ_804, 1 s
   "16_AQ_Data_R3_SPR_AQ_802" : Real = PLC "16_AQ_Data".R3_SPR_AQ_802, 1 s
   "80_From_HMI_MAN_AQ_INC_800" : Bool = PLC "80_From_HMI".MAN_AQ_INC_800, 1 s
   "80_From_HMI_MAN_AQ_DEC_806" : Bool = PLC "80_From_HMI".MAN_AQ_DEC_806, 1 s
   "80_From_HMI_MAN_AQ_INC_806" : Bool = PLC "80_From_HMI".MAN_AQ_INC_806, 1 s
   "80_From_HMI_MAN_AQ_DEC_804" : Bool = PLC "80_From_HMI".MAN_AQ_DEC_804, 1 s
   "80_From_HMI_MAN_AQ_INC_804" : Bool = PLC "80_From_HMI".MAN_AQ_INC_804, 1 s
   "80_From_HMI_MAN_AQ_DEC_802" : Bool = PLC "80_From_HMI".MAN_AQ_DEC_802, 1 s
   "80_From_HMI_MAN_AQ_INC_802" : Bool = PLC "80_From_HMI".MAN_AQ_INC_802, 1 s
   "80_From_HMI_MAN_AQ_DEC_800" : Bool = PLC "80_From_HMI".MAN_AQ_DEC_800, 1 s
   "86_Times_CV441_OPND_DLY" : Time = PLC "86_Times".CV441_OPND_DLY, 1 s
   "86_Times_CV401_OPND_DLY" : Time = PLC "86_Times".CV401_OPND_DLY, 1 s
   "86_Times_CV358_CLSD_DLY" : Time = PLC "86_Times".CV358_CLSD_DLY, 1 s
   "86_Times_CV341_CLSD_DLY" : Time = PLC "86_Times".CV341_CLSD_DLY, 1 s
   "86_Times_P305_STPD_DLY" : Time = PLC "86_Times".P305_STPD_DLY, 1 s
   "86_Times_P305_STRTD_DLY" : Time = PLC "86_Times".P305_STRTD_DLY, 1 s
   "86_Times_P304_STPD_DLY" : Time = PLC "86_Times".P304_STPD_DLY, 1 s
   "86_Times_P304_STRTD_DLY" : Time = PLC "86_Times".P304_STRTD_DLY, 1 s
   "86_Times_P303_STPD_DLY" : Time = PLC "86_Times".P303_STPD_DLY, 1 s
   "86_Times_CV407_MAX_TRVL_TIME" : Time = PLC "86_Times".CV407_MAX_TRVL_TIME, 1 s
   "86_Times_CV406_MAX_TRVL_TIME" : Time = PLC "86_Times".CV406_MAX_TRVL_TIME, 1 s
   "86_Times_CV358_MAX_TRVL_TIME" : Time = PLC "86_Times".CV358_MAX_TRVL_TIME, 1 s
   "86_Times_PIT416_TRGT_RMP_TIME" : Real = PLC "86_Times".PIT416_TRGT_RMP_TIME, 1 s
   "86_Times_CV441_MAX_TRVL_TIME" : Time = PLC "86_Times".CV441_MAX_TRVL_TIME, 1 s
   "86_Times_CV411_MAX_TRVL_TIME" : Time = PLC "86_Times".CV411_MAX_TRVL_TIME, 1 s
   "86_Times_CV341_MAX_TRVL_TIME" : Time = PLC "86_Times".CV341_MAX_TRVL_TIME, 1 s
   "86_Times_CV409_MAX_TRVL_TIME" : Time = PLC Alarms_Acknowledge.IGG_ALARM_ACKNLG_1, 1 s
   "86_Times_POST_FLUSH_DLY" : Time = PLC "86_Times".POST_FLUSH_DLY, 1 s
   "86_Times_GCU_FLUSH_TIME" : Time = PLC "86_Times".GCU_FLUSH_TIME, 1 s
   "86_Times_GCU_TNK_DRN_MAX_TIME" : Time = PLC "86_Times".GCU_TNK_DRN_MAX_TIME, 1 s
   "86_Times_CV341_OPND_DLY" : Time = PLC "86_Times".CV341_OPND_DLY, 1 s
   "86_Times_P303_STOP_TIME" : Time = PLC "86_Times".P303_STOP_TIME, 1 s
   "86_Times_E400_STOP_TIME" : Time = PLC "86_Times".E400_STOP_TIME, 1 s
   "86_Times_CV406_CLSD_DLY" : Time = PLC "86_Times".CV406_CLSD_DLY, 1 s
   "86_Times_CV405_OPND_DLY" : Time = PLC "86_Times".CV405_OPND_DLY, 1 s
   "86_Times_E400_RNG_DLY" : Time = PLC "86_Times".E400_RNG_DLY, 1 s
   "86_Times_E400_STRTD_DLY" : Time = PLC "86_Times".E400_STRTD_DLY, 1 s
   "86_Times_CV401_CLSD_DLY" : Time = PLC "86_Times".CV401_CLSD_DLY, 1 s
   "86_Times_CV441_CLSD_DLY" : Time = PLC "86_Times".CV441_CLSD_DLY, 1 s
   "86_Times_VLV_CNFG_DN_DLY" : Time = PLC "86_Times".VLV_CNFG_DN_DLY, 1 s
   "86_Times_P303_STRTD_DLY" : Time = PLC "86_Times".P303_STRTD_DLY, 1 s
   "86_Times_PRE_CV441_OPN_DLY" : Time = PLC "86_Times".PRE_CV441_OPN_DLY, 1 s
   "86_Times_GCU_TNK_FILL_MAX_TIME" : Time = PLC "86_Times".GCU_TNK_FILL_MAX_TIME, 1 s
   "86_Times_PRE_GCU_TNK_FILL_DLY" : Time = PLC "86_Times".PRE_GCU_TNK_FILL_DLY, 1 s
   "86_Times_STEP_MAX_TIME_STP_001" : Time = PLC "86_Times".STEP_MAX_TIME_STP_001, 1 s
   "86_Times_STEP_MAX_TIME_STP_005" : Time = PLC "86_Times".STEP_MAX_TIME_STP_005, 1 s
   "86_Times_STEP_MAX_TIME_STP_010" : Time = PLC "86_Times".STEP_MAX_TIME_STP_010, 1 s
   "86_Times_STEP_MAX_TIME_STP_020" : Time = PLC "86_Times".STEP_MAX_TIME_STP_020, 1 s
   "86_Times_STEP_MAX_TIME_STP_030" : Time = PLC "86_Times".STEP_MAX_TIME_STP_030, 1 s
   "86_Times_STEP_MAX_TIME_STP_040" : Time = PLC "86_Times".STEP_MAX_TIME_STP_040, 1 s
   "86_Times_STEP_MAX_TIME_STP_050" : Time = PLC "86_Times".STEP_MAX_TIME_STP_050, 1 s
   "86_Times_STEP_MAX_TIME_STP_060" : Time = PLC "86_Times".STEP_MAX_TIME_STP_060, 1 s
   "86_Times_STEP_MAX_TIME_STP_070" : Time = PLC "86_Times".STEP_MAX_TIME_STP_070, 1 s
   "86_Times_STEP_MAX_TIME_STP_080" : Time = PLC "86_Times".STEP_MAX_TIME_STP_080, 1 s
   "86_Times_STEP_MAX_TIME_STP_090" : Time = PLC "86_Times".STEP_MAX_TIME_STP_090, 1 s
   "86_Times_STEP_MAX_TIME_STP_100" : Time = PLC "86_Times".STEP_MAX_TIME_STP_100, 1 s
   "86_Times_STEP_MAX_TIME_STP_110" : Time = PLC "86_Times".STEP_MAX_TIME_STP_110, 1 s
   "86_Times_STEP_MAX_TIME_STP_120" : Time = PLC "86_Times".STEP_MAX_TIME_STP_120, 1 s
   "86_Times_STEP_MAX_TIME_STP_130" : Time = PLC "86_Times".STEP_MAX_TIME_STP_130, 1 s
   "86_Times_STEP_MAX_TIME_STP_140" : Time = PLC "86_Times".STEP_MAX_TIME_STP_140, 1 s
   "86_Times_STEP_MAX_TIME_STP_150" : Time = PLC "86_Times".STEP_MAX_TIME_STP_150, 1 s
   "86_Times_STEP_MAX_TIME_STP_160" : Time = PLC "86_Times".STEP_MAX_TIME_STP_160, 1 s
   "86_Times_STEP_MAX_TIME_STP_170" : Time = PLC "86_Times".STEP_MAX_TIME_STP_170, 1 s
   "86_Times_STEP_MAX_TIME_STP_180" : Time = PLC "86_Times".STEP_MAX_TIME_STP_180, 1 s
   "86_Times_STEP_MAX_TIME_STP_190" : Time = PLC "86_Times".STEP_MAX_TIME_STP_190, 1 s
   "86_Times_STEP_MAX_TIME_STP_200" : Time = PLC "86_Times".STEP_MAX_TIME_STP_200, 1 s
   "86_Times_STEP_MAX_TIME_STP_210" : Time = PLC "86_Times".STEP_MAX_TIME_STP_210, 1 s
   "86_Times_STEP_MAX_TIME_STP_220" : Time = PLC "86_Times".STEP_MAX_TIME_STP_220, 1 s
   "86_Times_STEP_MAX_TIME_STP_230" : Time = PLC "86_Times".STEP_MAX_TIME_STP_230, 1 s
   "86_Times_STEP_MAX_TIME_STP_240" : Time = PLC "86_Times".STEP_MAX_TIME_STP_240, 1 s
   "86_Times_STEP_MAX_TIME_STP_250" : Time = PLC "86_Times".STEP_MAX_TIME_STP_250, 1 s
   "86_Times_STEP_MAX_TIME_STP_260" : Time = PLC "86_Times".STEP_MAX_TIME_STP_260, 1 s
   "86_Times_STEP_MAX_TIME_STP_270" : Time = PLC "86_Times".STEP_MAX_TIME_STP_270, 1 s
   "86_Times_STEP_MAX_TIME_STP_280" : Time = PLC "86_Times".STEP_MAX_TIME_STP_280, 1 s
   "86_Times_STEP_MAX_TIME_STP_290" : Time = PLC "86_Times".STEP_MAX_TIME_STP_290, 1 s
   "86_Times_STEP_MAX_TIME_STP_300" : Time = PLC "86_Times".STEP_MAX_TIME_STP_300, 1 s
   "86_Times_STEP_MAX_TIME_STP_310" : Time = PLC "86_Times".STEP_MAX_TIME_STP_310, 1 s
   "86_Times_STEP_MAX_TIME_STP_320" : Time = PLC "86_Times".STEP_MAX_TIME_STP_320, 1 s
   "86_Times_STEP_MAX_TIME_STP_330" : Time = PLC "86_Times".STEP_MAX_TIME_STP_330, 1 s
   "86_Times_STEP_MAX_TIME_STP_340" : Time = PLC "86_Times".STEP_MAX_TIME_STP_340, 1 s
   "86_Times_STEP_MAX_TIME_STP_350" : Time = PLC "86_Times".STEP_MAX_TIME_STP_350, 1 s
   "86_Times_STEP_MAX_TIME_STP_360" : Time = PLC "86_Times".STEP_MAX_TIME_STP_360, 1 s
   "86_Times_STEP_MAX_TIME_STP_370" : Time = PLC "86_Times".STEP_MAX_TIME_STP_370, 1 s
   "86_Times_STEP_MAX_TIME_STP_380" : Time = PLC "86_Times".STEP_MAX_TIME_STP_380, 1 s
   "86_Times_STEP_MAX_TIME_STP_390" : Time = PLC "86_Times".STEP_MAX_TIME_STP_390, 1 s
   "86_Times_STEP_MAX_TIME_STP_400" : Time = PLC "86_Times".STEP_MAX_TIME_STP_400, 1 s
   "86_Times_STEP_MAX_TIME_STP_410" : Time = PLC "86_Times".STEP_MAX_TIME_STP_410, 1 s
   "86_Times_STEP_MAX_TIME_STP_420" : Time = PLC "86_Times".STEP_MAX_TIME_STP_420, 1 s
   "86_Times_STEP_MAX_TIME_STP_430" : Time = PLC "86_Times".STEP_MAX_TIME_STP_430, 1 s
   "86_Times_STEP_MAX_TIME_STP_440" : Time = PLC "86_Times".STEP_MAX_TIME_STP_440, 1 s
   "86_Times_STEP_MAX_TIME_STP_450" : Time = PLC "86_Times".STEP_MAX_TIME_STP_450, 1 s
   "86_Times_STEP_MAX_TIME_STP_460" : Time = PLC "86_Times".STEP_MAX_TIME_STP_460, 1 s
   "86_Times_STEP_MAX_TIME_STP_470" : Time = PLC "86_Times".STEP_MAX_TIME_STP_470, 1 s
   "86_Times_STEP_MAX_TIME_STP_480" : Time = PLC "86_Times".STEP_MAX_TIME_STP_480, 1 s
   "86_Times_STEP_MAX_TIME_STP_490" : Time = PLC "86_Times".STEP_MAX_TIME_STP_490, 1 s
   "86_Times_STEP_MAX_TIME_STP_500" : Time = PLC "86_Times".STEP_MAX_TIME_STP_500, 1 s
   "86_Times_STEP_MAX_TIME_STP_510" : Time = PLC "86_Times".STEP_MAX_TIME_STP_510, 1 s
   "86_Times_STEP_MAX_TIME_STP_520" : Time = PLC "86_Times".STEP_MAX_TIME_STP_520, 1 s
   "86_Times_STEP_MAX_TIME_STP_530" : Time = PLC "86_Times".STEP_MAX_TIME_STP_530, 1 s